REGION Network 15
   RUNG wire#powerrail
      { S7_Templates := "SrcType := Int" } EQ_Contact(in1 := "DB_general".Piston_2_Cursa_Completa, in2 := 25)
      R_Coil( "DB_HMI".Viz_Platforma_Libera )
   END_RUNG
   // the same network as SCL:
   IF "DB_general".Piston_2_Cursa_Completa = 25 THEN "DB_HMI".Viz_Platforma_Libera := FALSE; END_IF;
END_REGION
END_FUNCTION_BLOCK

FUNCTION_BLOCK "Piston_Incarcare"   // FB19, LAD
{ S7_Optimized_Access := 'FALSE' }
VERSION : 0.1
   VAR_TEMP   // added for the SCL form of the ladder/FBD networks
      _w1 : Bool;
      _w2 : Bool;
      _w3 : Bool;
      _w4 : Bool;
      _w5 : Bool;
      _w6 : Bool;
      _w7 : Bool;
   END_VAR
BEGIN

REGION Network 1
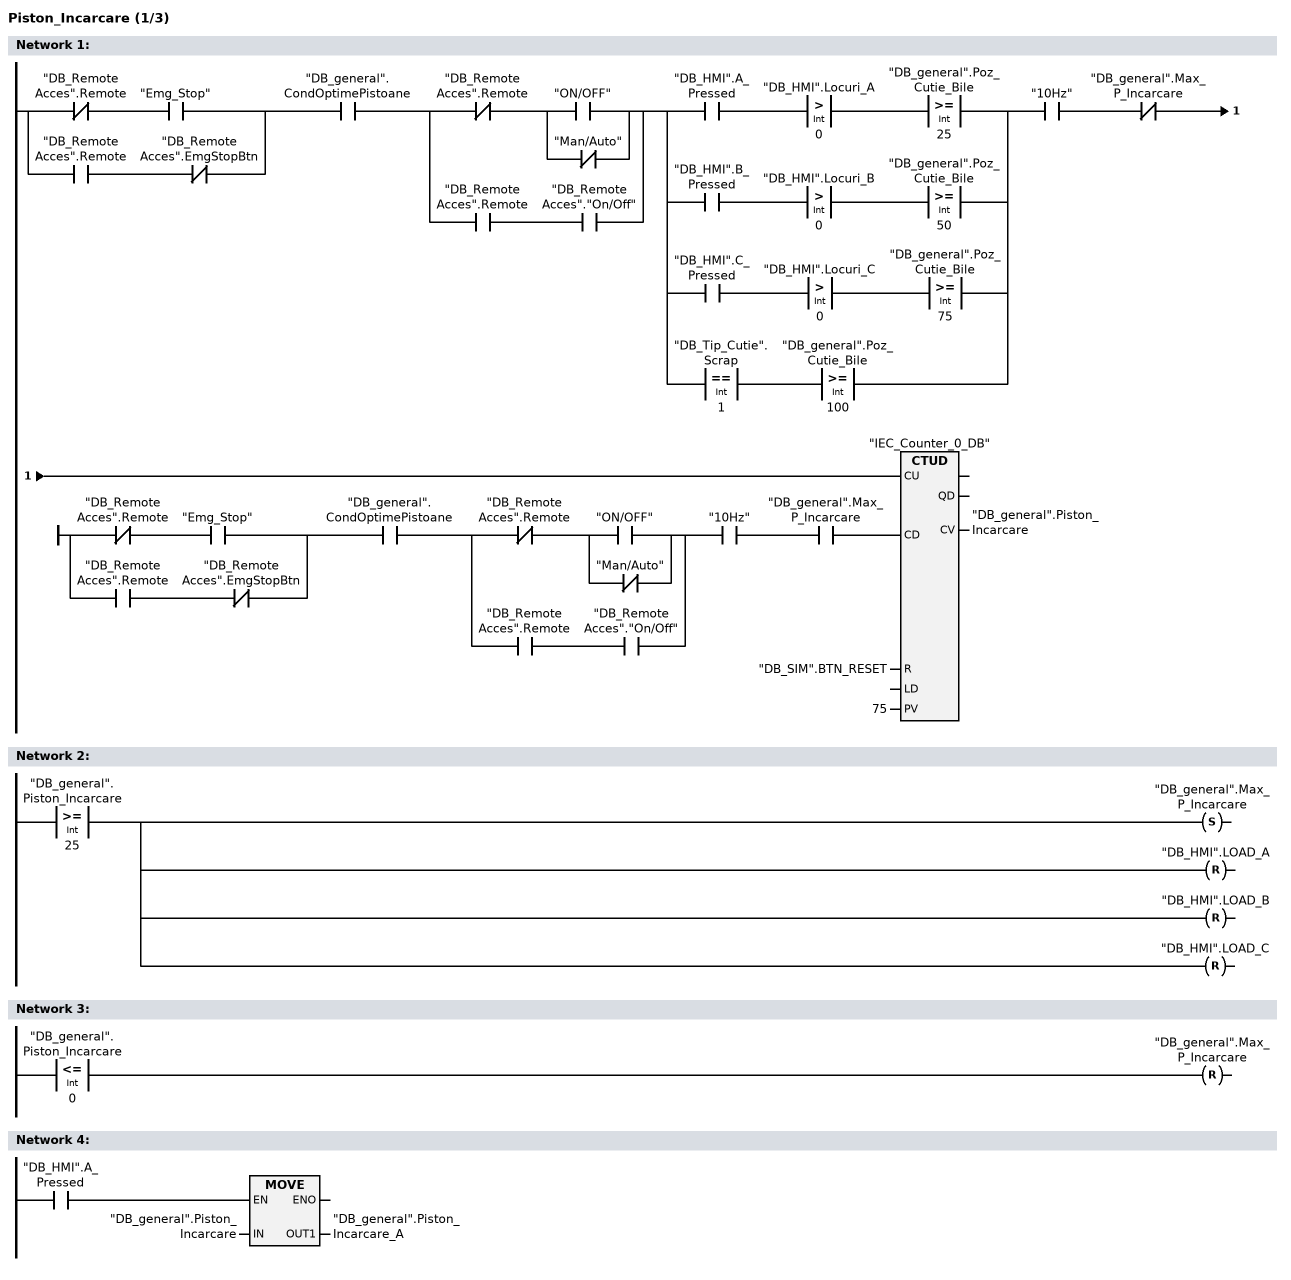
   "IEC_Counter_0_DB".CTUD(CU := ((NOT "DB_RemoteAcces".Remote AND "Emg_Stop") OR ("DB_RemoteAcces".Remote AND NOT "DB_RemoteAcces".EmgStopBtn)) AND "DB_general".CondOptimePistoane AND ((NOT "DB_RemoteAcces".Remote AND ("ON/OFF" OR NOT "Man/Auto")) OR ("DB_RemoteAcces".Remote AND "DB_RemoteAcces"."On/Off")) AND (("DB_HMI".A_Pressed AND ("DB_HMI".Locuri_A > 0) AND ("DB_general".Poz_Cutie_Bile >= 25)) OR ("DB_HMI".B_Pressed AND ("DB_HMI".Locuri_B > 0) AND ("DB_general".Poz_Cutie_Bile >= 50)) OR ("DB_HMI".C_Pressed AND ("DB_HMI".Locuri_C > 0) AND ("DB_general".Poz_Cutie_Bile >= 75)) OR (("DB_Tip_Cutie".Scrap = 1) AND ("DB_general".Poz_Cutie_Bile >= 100))) AND "10Hz" AND NOT "DB_general".Max_P_Incarcare,
                           CD := ((NOT "DB_RemoteAcces".Remote AND "Emg_Stop") OR ("DB_RemoteAcces".Remote AND NOT "DB_RemoteAcces".EmgStopBtn)) AND "DB_general".CondOptimePistoane AND ((NOT "DB_RemoteAcces".Remote AND ("ON/OFF" OR NOT "Man/Auto")) OR ("DB_RemoteAcces".Remote AND "DB_RemoteAcces"."On/Off")) AND "10Hz" AND "DB_general".Max_P_Incarcare,
                           R := "DB_SIM".BTN_RESET,
                           PV := 75,
                           CV => "DB_general".Piston_Incarcare);
END_REGION

REGION Network 2
   RUNG wire#powerrail
      { S7_Templates := "SrcType := Int" } GE_Contact(in1 := "DB_general".Piston_Incarcare, in2 := 25)
      wire#w1
      S_Coil( "DB_general".Max_P_Incarcare )
   END_RUNG
   RUNG wire#w1
      R_Coil( "DB_HMI".LOAD_A )
   END_RUNG
   RUNG wire#w1
      R_Coil( "DB_HMI".LOAD_B )
   END_RUNG
   RUNG wire#w1
      R_Coil( "DB_HMI".LOAD_C )
   END_RUNG
   // the same network as SCL:
   IF "DB_general".Piston_Incarcare >= 25 THEN
       "DB_general".Max_P_Incarcare := TRUE;
       "DB_HMI".LOAD_A := FALSE;
       "DB_HMI".LOAD_B := FALSE;
       "DB_HMI".LOAD_C := FALSE;
   END_IF;
END_REGION

REGION Network 3
   RUNG wire#powerrail
      { S7_Templates := "SrcType := Int" } LE_Contact(in1 := "DB_general".Piston_Incarcare, in2 := 0)
      R_Coil( "DB_general".Max_P_Incarcare )
   END_RUNG
   // the same network as SCL:
   IF "DB_general".Piston_Incarcare <= 0 THEN "DB_general".Max_P_Incarcare := FALSE; END_IF;
END_REGION

REGION Network 4
   RUNG wire#powerrail
      Contact( "DB_HMI".A_Pressed )
      { S7_GenerateENO := "TRUE" } Move(in := "DB_general".Piston_Incarcare, out1 => "DB_general".Piston_Incarcare_A)
   END_RUNG
   // the same network as SCL:
   IF "DB_HMI".A_Pressed THEN "DB_general".Piston_Incarcare_A := "DB_general".Piston_Incarcare; END_IF;
END_REGION

REGION Network 5
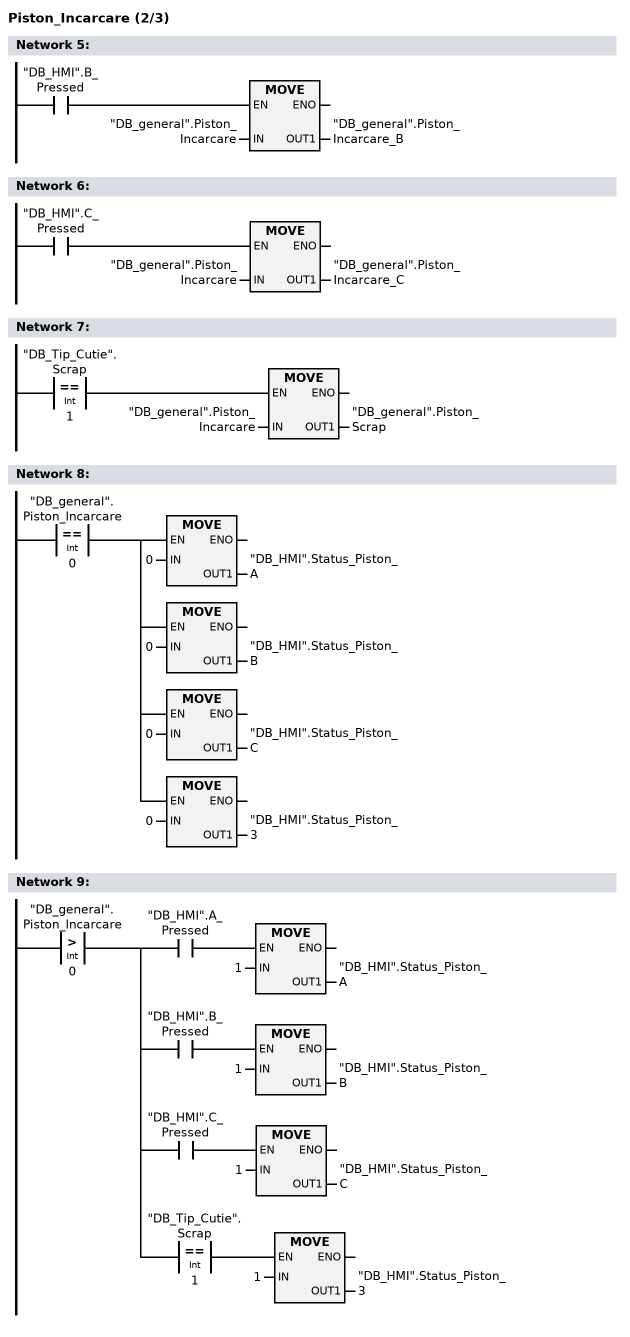
   RUNG wire#powerrail
      Contact( "DB_HMI".B_Pressed )
      { S7_GenerateENO := "TRUE" } Move(in := "DB_general".Piston_Incarcare, out1 => "DB_general".Piston_Incarcare_B)
   END_RUNG
   // the same network as SCL:
   IF "DB_HMI".B_Pressed THEN "DB_general".Piston_Incarcare_B := "DB_general".Piston_Incarcare; END_IF;
END_REGION

REGION Network 6
   RUNG wire#powerrail
      Contact( "DB_HMI".C_Pressed )
      { S7_GenerateENO := "TRUE" } Move(in := "DB_general".Piston_Incarcare, out1 => "DB_general".Piston_Incarcare_C)
   END_RUNG
   // the same network as SCL:
   IF "DB_HMI".C_Pressed THEN "DB_general".Piston_Incarcare_C := "DB_general".Piston_Incarcare; END_IF;
END_REGION

REGION Network 7
   RUNG wire#powerrail
      { S7_Templates := "SrcType := Int" } EQ_Contact(in1 := "DB_Tip_Cutie".Scrap, in2 := 1)
      { S7_GenerateENO := "TRUE" } Move(in := "DB_general".Piston_Incarcare, out1 => "DB_general".Piston_Scrap)
   END_RUNG
   // the same network as SCL:
   IF "DB_Tip_Cutie".Scrap = 1 THEN "DB_general".Piston_Scrap := "DB_general".Piston_Incarcare; END_IF;
END_REGION

REGION Network 8
   RUNG wire#powerrail
      { S7_Templates := "SrcType := Int" } EQ_Contact(in1 := "DB_general".Piston_Incarcare, in2 := 0)
      wire#w1
      { S7_GenerateENO := "TRUE" } Move(in := 0, out1 => "DB_HMI".Status_Piston_A)
   END_RUNG
   RUNG wire#w1
      { S7_GenerateENO := "TRUE" } Move(in := 0, out1 => "DB_HMI".Status_Piston_B)
   END_RUNG
   RUNG wire#w1
      { S7_GenerateENO := "TRUE" } Move(in := 0, out1 => "DB_HMI".Status_Piston_C)
   END_RUNG
   RUNG wire#w1
      { S7_GenerateENO := "TRUE" } Move(in := 0, out1 => "DB_HMI".Status_Piston_3)
   END_RUNG
   // the same network as SCL:
   IF "DB_general".Piston_Incarcare = 0 THEN
       "DB_HMI".Status_Piston_A := 0;
       "DB_HMI".Status_Piston_B := 0;
       "DB_HMI".Status_Piston_C := 0;
       "DB_HMI".Status_Piston_3 := 0;
   END_IF;
END_REGION

REGION Network 9
   RUNG wire#powerrail
      { S7_Templates := "SrcType := Int" } GT_Contact(in1 := "DB_general".Piston_Incarcare, in2 := 0)
      wire#w1
      Contact( "DB_HMI".A_Pressed )
      { S7_GenerateENO := "TRUE" } Move(in := 1, out1 => "DB_HMI".Status_Piston_A)
   END_RUNG
   RUNG wire#w1
      Contact( "DB_HMI".B_Pressed )
      { S7_GenerateENO := "TRUE" } Move(in := 1, out1 => "DB_HMI".Status_Piston_B)
   END_RUNG
   RUNG wire#w1
      Contact( "DB_HMI".C_Pressed )
      { S7_GenerateENO := "TRUE" } Move(in := 1, out1 => "DB_HMI".Status_Piston_C)
   END_RUNG
   RUNG wire#w1
      { S7_Templates := "SrcType := Int" } EQ_Contact(in1 := "DB_Tip_Cutie".Scrap, in2 := 1)
      { S7_GenerateENO := "TRUE" } Move(in := 1, out1 => "DB_HMI".Status_Piston_3)
   END_RUNG
   // the same network as SCL:
   #_w1 := "DB_general".Piston_Incarcare > 0;
   IF #_w1 AND "DB_HMI".A_Pressed THEN "DB_HMI".Status_Piston_A := 1; END_IF;
   IF #_w1 AND "DB_HMI".B_Pressed THEN "DB_HMI".Status_Piston_B := 1; END_IF;
   IF #_w1 AND "DB_HMI".C_Pressed THEN "DB_HMI".Status_Piston_C := 1; END_IF;
   IF #_w1 AND ("DB_Tip_Cutie".Scrap = 1) THEN "DB_HMI".Status_Piston_3 := 1; END_IF;
END_REGION

REGION Network 10
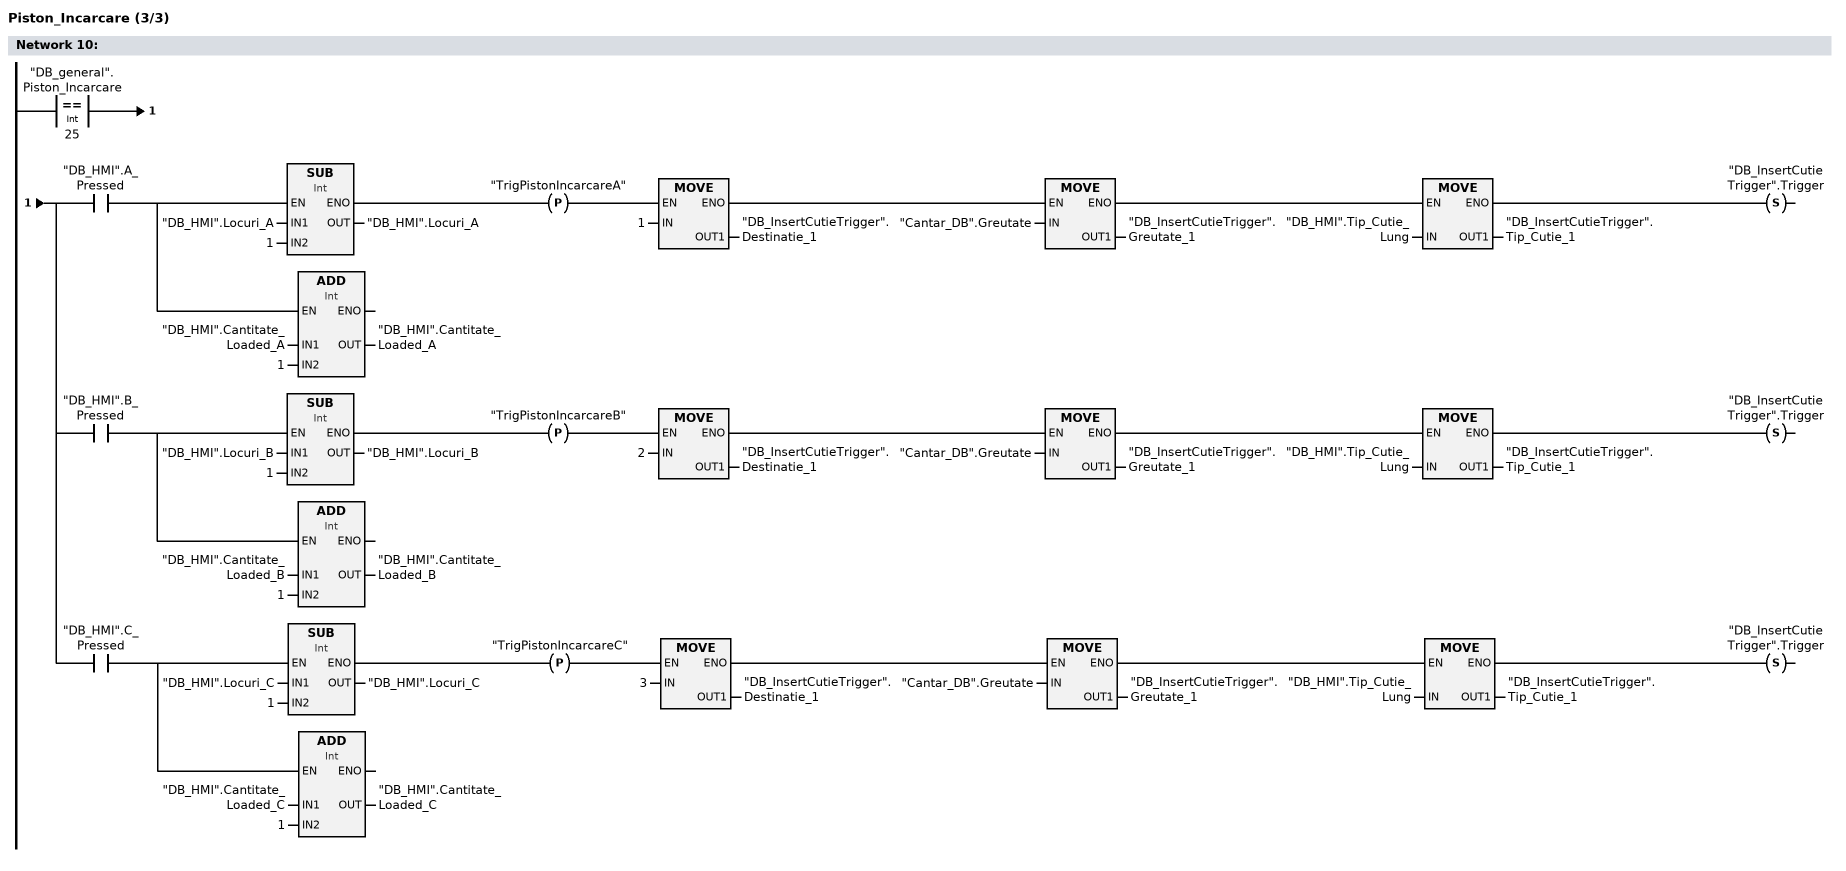
   RUNG wire#powerrail
      { S7_Templates := "SrcType := Int" } EQ_Contact(in1 := "DB_general".Piston_Incarcare, in2 := 25)
      wire#w1
      Contact( "DB_HMI".A_Pressed )
      wire#w2
      { S7_Templates := "SrcType := Int"; S7_GenerateENO := "TRUE" } Sub(in1 := "DB_HMI".Locuri_A, in2 := 1, out => "DB_HMI".Locuri_A)
      P_Trig( "TrigPistonIncarcareA" )
      { S7_GenerateENO := "TRUE" } Move(in := 1, out1 => "DB_InsertCutieTrigger".Destinatie_1)
      { S7_GenerateENO := "TRUE" } Move(in := "Cantar_DB".Greutate, out1 => "DB_InsertCutieTrigger".Greutate_1)
      { S7_GenerateENO := "TRUE" } Move(in := "DB_HMI".Tip_Cutie_Lung, out1 => "DB_InsertCutieTrigger".Tip_Cutie_1)
      S_Coil( "DB_InsertCutieTrigger".Trigger )
   END_RUNG
   RUNG wire#w2
      { S7_Templates := "SrcType := Int"; S7_GenerateENO := "TRUE" } Add(in1 := "DB_HMI".Cantitate_Loaded_A, in2 := 1, out => "DB_HMI".Cantitate_Loaded_A)
   END_RUNG
   RUNG wire#w1
      Contact( "DB_HMI".B_Pressed )
      wire#w3
      { S7_Templates := "SrcType := Int"; S7_GenerateENO := "TRUE" } Sub(in1 := "DB_HMI".Locuri_B, in2 := 1, out => "DB_HMI".Locuri_B)
      P_Trig( "TrigPistonIncarcareB" )
      { S7_GenerateENO := "TRUE" } Move(in := 2, out1 => "DB_InsertCutieTrigger".Destinatie_1)
      { S7_GenerateENO := "TRUE" } Move(in := "Cantar_DB".Greutate, out1 => "DB_InsertCutieTrigger".Greutate_1)
      { S7_GenerateENO := "TRUE" } Move(in := "DB_HMI".Tip_Cutie_Lung, out1 => "DB_InsertCutieTrigger".Tip_Cutie_1)
      S_Coil( "DB_InsertCutieTrigger".Trigger )
   END_RUNG
   RUNG wire#w3
      { S7_Templates := "SrcType := Int"; S7_GenerateENO := "TRUE" } Add(in1 := "DB_HMI".Cantitate_Loaded_B, in2 := 1, out => "DB_HMI".Cantitate_Loaded_B)
   END_RUNG
   RUNG wire#w1
      Contact( "DB_HMI".C_Pressed )
      wire#w4
      { S7_Templates := "SrcType := Int"; S7_GenerateENO := "TRUE" } Sub(in1 := "DB_HMI".Locuri_C, in2 := 1, out => "DB_HMI".Locuri_C)
      P_Trig( "TrigPistonIncarcareC" )
      { S7_GenerateENO := "TRUE" } Move(in := 3, out1 => "DB_InsertCutieTrigger".Destinatie_1)
      { S7_GenerateENO := "TRUE" } Move(in := "Cantar_DB".Greutate, out1 => "DB_InsertCutieTrigger".Greutate_1)
      { S7_GenerateENO := "TRUE" } Move(in := "DB_HMI".Tip_Cutie_Lung, out1 => "DB_InsertCutieTrigger".Tip_Cutie_1)
      S_Coil( "DB_InsertCutieTrigger".Trigger )
   END_RUNG
   RUNG wire#w4
      { S7_Templates := "SrcType := Int"; S7_GenerateENO := "TRUE" } Add(in1 := "DB_HMI".Cantitate_Loaded_C, in2 := 1, out => "DB_HMI".Cantitate_Loaded_C)
   END_RUNG
   // the same network as SCL:
   // ENO of a box is taken as its EN; it also drops when the box reports an error
   #_w1 := "DB_general".Piston_Incarcare = 25;
   #_w2 := #_w1 AND "DB_HMI".A_Pressed;
   IF #_w2 THEN "DB_HMI".Locuri_A := "DB_HMI".Locuri_A - 1; END_IF;
   #_w3 := #_w2 AND NOT "TrigPistonIncarcareA";   // rising edge
   "TrigPistonIncarcareA" := #_w2;
   IF #_w3 THEN
       "DB_InsertCutieTrigger".Destinatie_1 := 1;
       "DB_InsertCutieTrigger".Greutate_1 := "Cantar_DB".Greutate;
       "DB_InsertCutieTrigger".Tip_Cutie_1 := "DB_HMI".Tip_Cutie_Lung;
       "DB_InsertCutieTrigger".Trigger := TRUE;
   END_IF;
   IF #_w2 THEN "DB_HMI".Cantitate_Loaded_A := "DB_HMI".Cantitate_Loaded_A + 1; END_IF;
   #_w4 := #_w1 AND "DB_HMI".B_Pressed;
   IF #_w4 THEN "DB_HMI".Locuri_B := "DB_HMI".Locuri_B - 1; END_IF;
   #_w5 := #_w4 AND NOT "TrigPistonIncarcareB";   // rising edge
   "TrigPistonIncarcareB" := #_w4;
   IF #_w5 THEN
       "DB_InsertCutieTrigger".Destinatie_1 := 2;
       "DB_InsertCutieTrigger".Greutate_1 := "Cantar_DB".Greutate;
       "DB_InsertCutieTrigger".Tip_Cutie_1 := "DB_HMI".Tip_Cutie_Lung;
       "DB_InsertCutieTrigger".Trigger := TRUE;
   END_IF;
   IF #_w4 THEN "DB_HMI".Cantitate_Loaded_B := "DB_HMI".Cantitate_Loaded_B + 1; END_IF;
   #_w6 := #_w1 AND "DB_HMI".C_Pressed;
   IF #_w6 THEN "DB_HMI".Locuri_C := "DB_HMI".Locuri_C - 1; END_IF;
   #_w7 := #_w6 AND NOT "TrigPistonIncarcareC";   // rising edge
   "TrigPistonIncarcareC" := #_w6;
   IF #_w7 THEN
       "DB_InsertCutieTrigger".Destinatie_1 := 3;
       "DB_InsertCutieTrigger".Greutate_1 := "Cantar_DB".Greutate;
       "DB_InsertCutieTrigger".Tip_Cutie_1 := "DB_HMI".Tip_Cutie_Lung;
       "DB_InsertCutieTrigger".Trigger := TRUE;
   END_IF;
   IF #_w6 THEN "DB_HMI".Cantitate_Loaded_C := "DB_HMI".Cantitate_Loaded_C + 1; END_IF;
END_REGION
END_FUNCTION_BLOCK

FUNCTION "Vizibilitate_Platforme/Colete" : Void   // FC1, LAD
{ S7_Optimized_Access := 'FALSE' }
VERSION : 0.1
BEGIN

REGION Network 1: Caz A apasat setare vizibilitate / Sichtbarkeitseinstellung für Fall „A“.
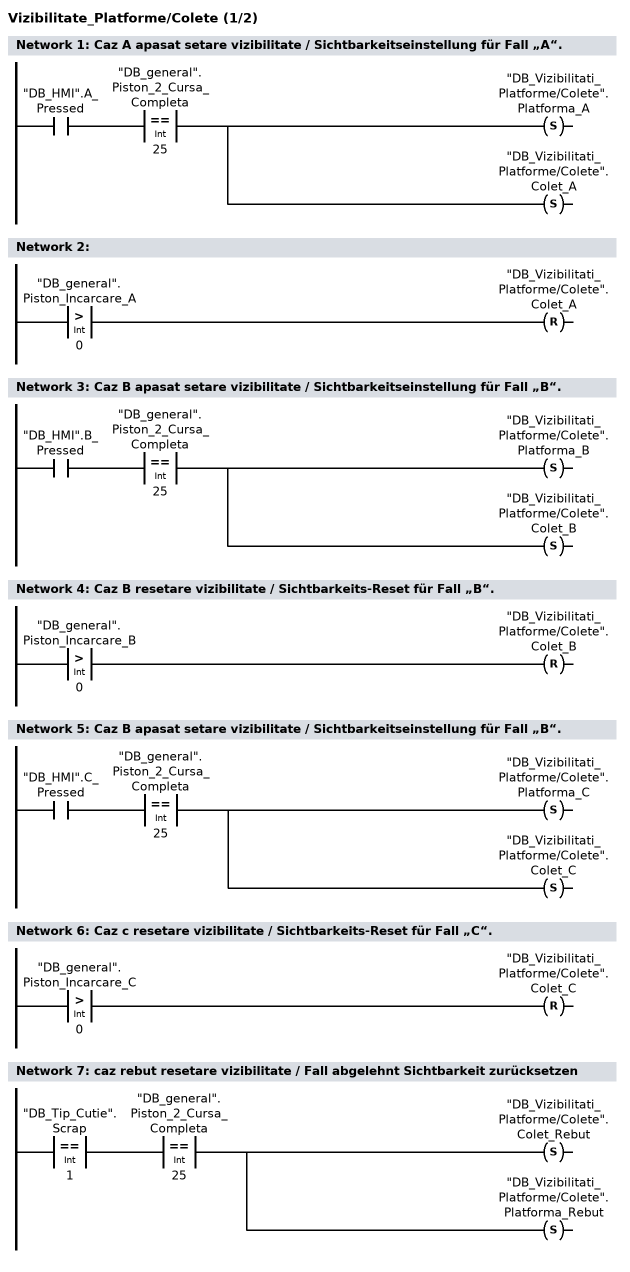
   RUNG wire#powerrail
      Contact( "DB_HMI".A_Pressed )
      { S7_Templates := "SrcType := Int" } EQ_Contact(in1 := "DB_general".Piston_2_Cursa_Completa, in2 := 25)
      wire#w1
      S_Coil( "DB_Vizibilitati_Platforme/Colete".Platforma_A )
   END_RUNG
   RUNG wire#w1
      S_Coil( "DB_Vizibilitati_Platforme/Colete".Colet_A )
   END_RUNG
   // the same network as SCL:
   IF "DB_HMI".A_Pressed AND ("DB_general".Piston_2_Cursa_Completa = 25) THEN
       "DB_Vizibilitati_Platforme/Colete".Platforma_A := TRUE;
       "DB_Vizibilitati_Platforme/Colete".Colet_A := TRUE;
   END_IF;
END_REGION

REGION Network 2
   RUNG wire#powerrail
      { S7_Templates := "SrcType := Int" } GT_Contact(in1 := "DB_general".Piston_Incarcare_A, in2 := 0)
      R_Coil( "DB_Vizibilitati_Platforme/Colete".Colet_A )
   END_RUNG
   // the same network as SCL:
   IF "DB_general".Piston_Incarcare_A > 0 THEN "DB_Vizibilitati_Platforme/Colete".Colet_A := FALSE; END_IF;
END_REGION

REGION Network 3: Caz B apasat setare vizibilitate / Sichtbarkeitseinstellung für Fall „B“.
   RUNG wire#powerrail
      Contact( "DB_HMI".B_Pressed )
      { S7_Templates := "SrcType := Int" } EQ_Contact(in1 := "DB_general".Piston_2_Cursa_Completa, in2 := 25)
      wire#w1
      S_Coil( "DB_Vizibilitati_Platforme/Colete".Platforma_B )
   END_RUNG
   RUNG wire#w1
      S_Coil( "DB_Vizibilitati_Platforme/Colete".Colet_B )
   END_RUNG
   // the same network as SCL:
   IF "DB_HMI".B_Pressed AND ("DB_general".Piston_2_Cursa_Completa = 25) THEN
       "DB_Vizibilitati_Platforme/Colete".Platforma_B := TRUE;
       "DB_Vizibilitati_Platforme/Colete".Colet_B := TRUE;
   END_IF;
END_REGION

REGION Network 4: Caz B resetare vizibilitate / Sichtbarkeits-Reset für Fall „B“.
   RUNG wire#powerrail
      { S7_Templates := "SrcType := Int" } GT_Contact(in1 := "DB_general".Piston_Incarcare_B, in2 := 0)
      R_Coil( "DB_Vizibilitati_Platforme/Colete".Colet_B )
   END_RUNG
   // the same network as SCL:
   IF "DB_general".Piston_Incarcare_B > 0 THEN "DB_Vizibilitati_Platforme/Colete".Colet_B := FALSE; END_IF;
END_REGION

REGION Network 5: Caz B apasat setare vizibilitate / Sichtbarkeitseinstellung für Fall „B“.
   RUNG wire#powerrail
      Contact( "DB_HMI".C_Pressed )
      { S7_Templates := "SrcType := Int" } EQ_Contact(in1 := "DB_general".Piston_2_Cursa_Completa, in2 := 25)
      wire#w1
      S_Coil( "DB_Vizibilitati_Platforme/Colete".Platforma_C )
   END_RUNG
   RUNG wire#w1
      S_Coil( "DB_Vizibilitati_Platforme/Colete".Colet_C )
   END_RUNG
   // the same network as SCL:
   IF "DB_HMI".C_Pressed AND ("DB_general".Piston_2_Cursa_Completa = 25) THEN
       "DB_Vizibilitati_Platforme/Colete".Platforma_C := TRUE;
       "DB_Vizibilitati_Platforme/Colete".Colet_C := TRUE;
   END_IF;
END_REGION

REGION Network 6: Caz c resetare vizibilitate / Sichtbarkeits-Reset für Fall „C“.
   RUNG wire#powerrail
      { S7_Templates := "SrcType := Int" } GT_Contact(in1 := "DB_general".Piston_Incarcare_C, in2 := 0)
      R_Coil( "DB_Vizibilitati_Platforme/Colete".Colet_C )
   END_RUNG
   // the same network as SCL:
   IF "DB_general".Piston_Incarcare_C > 0 THEN "DB_Vizibilitati_Platforme/Colete".Colet_C := FALSE; END_IF;
END_REGION

REGION Network 7: caz rebut resetare vizibilitate / Fall abgelehnt Sichtbarkeit zurücksetzen
   RUNG wire#powerrail
      { S7_Templates := "SrcType := Int" } EQ_Contact(in1 := "DB_Tip_Cutie".Scrap, in2 := 1)
      { S7_Templates := "SrcType := Int" } EQ_Contact(in1 := "DB_general".Piston_2_Cursa_Completa, in2 := 25)
      wire#w1
      S_Coil( "DB_Vizibilitati_Platforme/Colete".Colet_Rebut )
   END_RUNG
   RUNG wire#w1
      S_Coil( "DB_Vizibilitati_Platforme/Colete".Platforma_Rebut )
   END_RUNG
   // the same network as SCL:
   IF ("DB_Tip_Cutie".Scrap = 1) AND ("DB_general".Piston_2_Cursa_Completa = 25) THEN
       "DB_Vizibilitati_Platforme/Colete".Colet_Rebut := TRUE;
       "DB_Vizibilitati_Platforme/Colete".Platforma_Rebut := TRUE;
   END_IF;
END_REGION

REGION Network 8
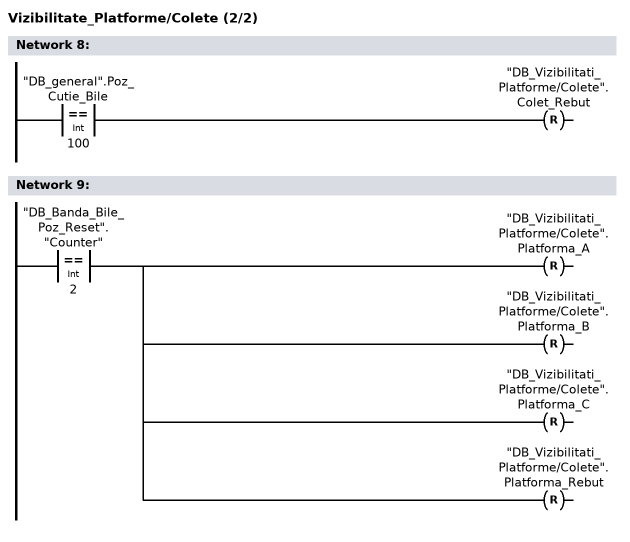
   RUNG wire#powerrail
      { S7_Templates := "SrcType := Int" } EQ_Contact(in1 := "DB_general".Poz_Cutie_Bile, in2 := 100)
      R_Coil( "DB_Vizibilitati_Platforme/Colete".Colet_Rebut )
   END_RUNG
   // the same network as SCL:
   IF "DB_general".Poz_Cutie_Bile = 100 THEN "DB_Vizibilitati_Platforme/Colete".Colet_Rebut := FALSE; END_IF;
END_REGION

REGION Network 9
   RUNG wire#powerrail
      { S7_Templates := "SrcType := Int" } EQ_Contact(in1 := "DB_Banda_Bile_Poz_Reset"."Counter", in2 := 2)
      wire#w1
      R_Coil( "DB_Vizibilitati_Platforme/Colete".Platforma_A )
   END_RUNG
   RUNG wire#w1
      R_Coil( "DB_Vizibilitati_Platforme/Colete".Platforma_B )
   END_RUNG
   RUNG wire#w1
      R_Coil( "DB_Vizibilitati_Platforme/Colete".Platforma_C )
   END_RUNG
   RUNG wire#w1
      R_Coil( "DB_Vizibilitati_Platforme/Colete".Platforma_Rebut )
   END_RUNG
   // the same network as SCL:
   IF "DB_Banda_Bile_Poz_Reset"."Counter" = 2 THEN
       "DB_Vizibilitati_Platforme/Colete".Platforma_A := FALSE;
       "DB_Vizibilitati_Platforme/Colete".Platforma_B := FALSE;
       "DB_Vizibilitati_Platforme/Colete".Platforma_C := FALSE;
       "DB_Vizibilitati_Platforme/Colete".Platforma_Rebut := FALSE;
   END_IF;
END_REGION
END_FUNCTION

// folder: Statie Incarcare/Functii

FUNCTION_BLOCK "Banda_Bile"   // FB16, SCL
{ S7_Optimized_Access := 'FALSE' }
VERSION : 0.1
   VAR_INPUT
      "Man/Auto" : Bool;
      BTN_Transport : Bool;
      Poz_Cutie_1 : Int;
      Emg_Stop : Bool;
      Btn_A : Bool;
      Btn_B : Bool;
      Btn_C : Bool;
   END_VAR
   VAR_OUTPUT
      Status_Banda_Bile : Bool;
   END_VAR
   VAR
      Btn_Transport_Pressed : Bool;
   END_VAR
BEGIN
   //IF #BTN_Transport THEN
     //  #Btn_Transport_Pressed := true;

   //END_IF;



       IF #Poz_Cutie_1 >48 AND "DB_HMI".Transport AND "DB_general".Piston_2_Cursa_Completa =0 AND (#Btn_A OR #Btn_B OR #Btn_C OR "DB_Tip_Cutie".Scrap = 1) THEN

           #Status_Banda_Bile := TRUE;
       ELSE
           #Status_Banda_Bile := FALSE;
           #Btn_Transport_Pressed := FALSE;


       END_IF;
END_FUNCTION_BLOCK

FUNCTION "Banda_Bile_Poz_Reset" : Void   // FC9, LAD
{ S7_Optimized_Access := 'FALSE' }
VERSION : 0.1
BEGIN

REGION Network 1
   // Atunci cand platforma cu bile trece de doua ori prin dreptul unui punct inseamna ca s a efectuat descarcarea si ca op ar trebui sa introduca o alta destinatie
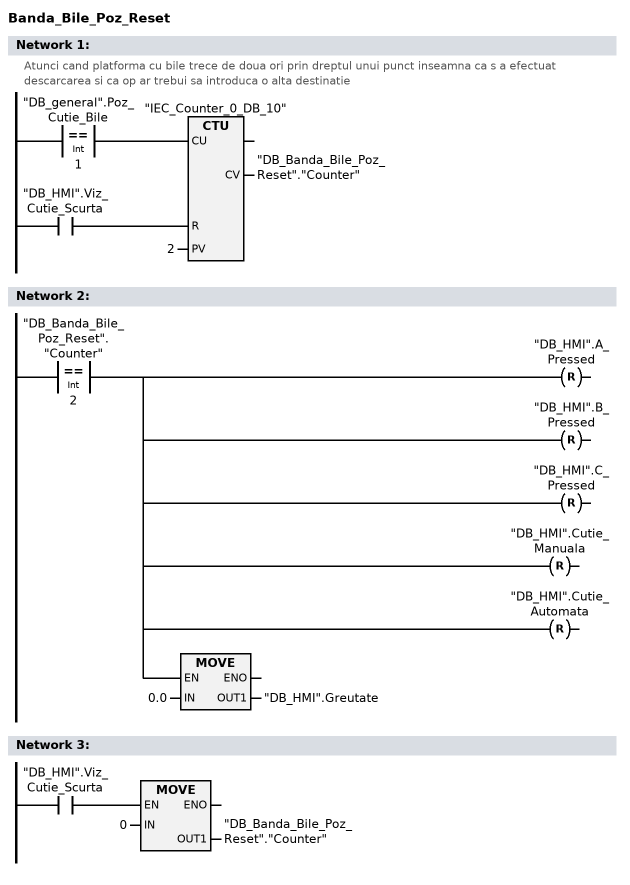
   "IEC_Counter_0_DB_10".CTU(CU := "DB_general".Poz_Cutie_Bile = 1,
                           R := "DB_HMI".Viz_Cutie_Scurta,
                           PV := 2,
                           CV => "DB_Banda_Bile_Poz_Reset"."Counter");
END_REGION

REGION Network 2
   RUNG wire#powerrail
      { S7_Templates := "SrcType := Int" } EQ_Contact(in1 := "DB_Banda_Bile_Poz_Reset"."Counter", in2 := 2)
      wire#w1
      R_Coil( "DB_HMI".A_Pressed )
   END_RUNG
   RUNG wire#w1
      R_Coil( "DB_HMI".B_Pressed )
   END_RUNG
   RUNG wire#w1
      R_Coil( "DB_HMI".C_Pressed )
   END_RUNG
   RUNG wire#w1
      R_Coil( "DB_HMI".Cutie_Manuala )
   END_RUNG
   RUNG wire#w1
      R_Coil( "DB_HMI".Cutie_Automata )
   END_RUNG
   RUNG wire#w1
      { S7_GenerateENO := "TRUE" } Move(in := 0.0, out1 => "DB_HMI".Greutate)
   END_RUNG
   // the same network as SCL:
   IF "DB_Banda_Bile_Poz_Reset"."Counter" = 2 THEN
       "DB_HMI".A_Pressed := FALSE;
       "DB_HMI".B_Pressed := FALSE;
       "DB_HMI".C_Pressed := FALSE;
       "DB_HMI".Cutie_Manuala := FALSE;
       "DB_HMI".Cutie_Automata := FALSE;
       "DB_HMI".Greutate := 0.0;
   END_IF;
END_REGION

REGION Network 3
   RUNG wire#powerrail
      Contact( "DB_HMI".Viz_Cutie_Scurta )
      { S7_GenerateENO := "TRUE" } Move(in := 0, out1 => "DB_Banda_Bile_Poz_Reset"."Counter")
   END_RUNG
   // the same network as SCL:
   IF "DB_HMI".Viz_Cutie_Scurta THEN "DB_Banda_Bile_Poz_Reset"."Counter" := 0; END_IF;
END_REGION
END_FUNCTION

FUNCTION "GreutateTotala" : Void   // FC14, LAD
{ S7_Optimized_Access := 'FALSE' }
VERSION : 0.1
BEGIN

REGION Network 1
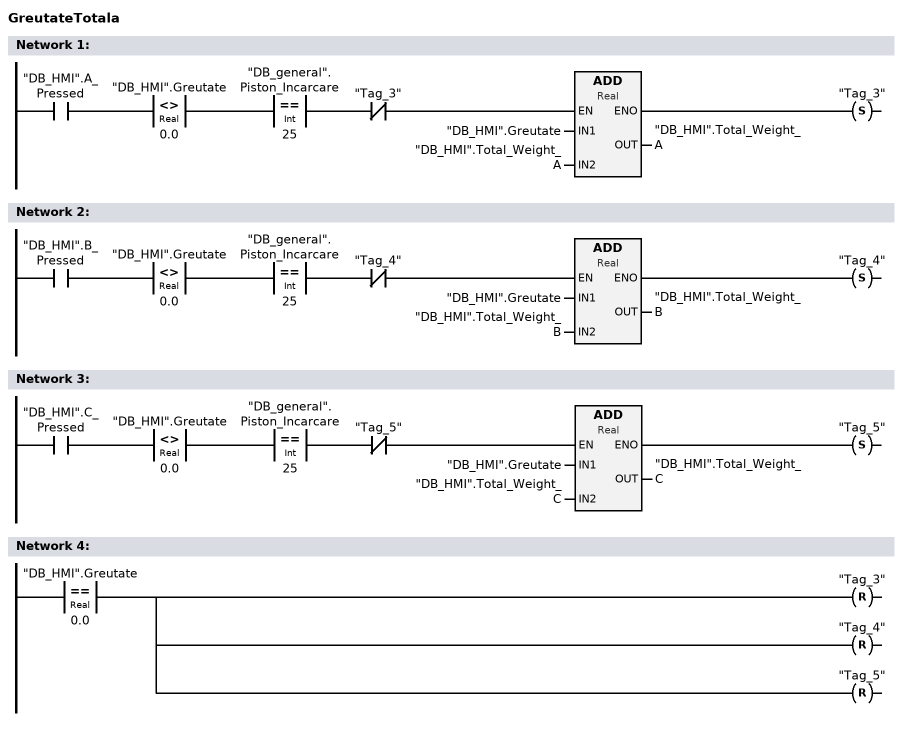
   RUNG wire#powerrail
      Contact( "DB_HMI".A_Pressed )
      { S7_Templates := "SrcType := Real" } NE_Contact(in1 := "DB_HMI".Greutate, in2 := 0.0)
      { S7_Templates := "SrcType := Int" } EQ_Contact(in1 := "DB_general".Piston_Incarcare, in2 := 25)
      I_Contact( "Tag_3" )
      { S7_Templates := "SrcType := Real"; S7_GenerateENO := "TRUE" } Add(in1 := "DB_HMI".Greutate, in2 := "DB_HMI".Total_Weight_A, out => "DB_HMI".Total_Weight_A)
      S_Coil( "Tag_3" )
   END_RUNG
   // the same network as SCL:
   // ENO of a box is taken as its EN; it also drops when the box reports an error
   IF "DB_HMI".A_Pressed AND ("DB_HMI".Greutate <> 0.0) AND ("DB_general".Piston_Incarcare = 25) AND NOT "Tag_3" THEN
       "DB_HMI".Total_Weight_A := "DB_HMI".Greutate + "DB_HMI".Total_Weight_A;
       "Tag_3" := TRUE;
   END_IF;
END_REGION

REGION Network 2
   RUNG wire#powerrail
      Contact( "DB_HMI".B_Pressed )
      { S7_Templates := "SrcType := Real" } NE_Contact(in1 := "DB_HMI".Greutate, in2 := 0.0)
      { S7_Templates := "SrcType := Int" } EQ_Contact(in1 := "DB_general".Piston_Incarcare, in2 := 25)
      I_Contact( "Tag_4" )
      { S7_Templates := "SrcType := Real"; S7_GenerateENO := "TRUE" } Add(in1 := "DB_HMI".Greutate, in2 := "DB_HMI".Total_Weight_B, out => "DB_HMI".Total_Weight_B)
      S_Coil( "Tag_4" )
   END_RUNG
   // the same network as SCL:
   // ENO of a box is taken as its EN; it also drops when the box reports an error
   IF "DB_HMI".B_Pressed AND ("DB_HMI".Greutate <> 0.0) AND ("DB_general".Piston_Incarcare = 25) AND NOT "Tag_4" THEN
       "DB_HMI".Total_Weight_B := "DB_HMI".Greutate + "DB_HMI".Total_Weight_B;
       "Tag_4" := TRUE;
   END_IF;
END_REGION

REGION Network 3
   RUNG wire#powerrail
      Contact( "DB_HMI".C_Pressed )
      { S7_Templates := "SrcType := Real" } NE_Contact(in1 := "DB_HMI".Greutate, in2 := 0.0)
      { S7_Templates := "SrcType := Int" } EQ_Contact(in1 := "DB_general".Piston_Incarcare, in2 := 25)
      I_Contact( "Tag_5" )
      { S7_Templates := "SrcType := Real"; S7_GenerateENO := "TRUE" } Add(in1 := "DB_HMI".Greutate, in2 := "DB_HMI".Total_Weight_C, out => "DB_HMI".Total_Weight_C)
      S_Coil( "Tag_5" )
   END_RUNG
   // the same network as SCL:
   // ENO of a box is taken as its EN; it also drops when the box reports an error
   IF "DB_HMI".C_Pressed AND ("DB_HMI".Greutate <> 0.0) AND ("DB_general".Piston_Incarcare = 25) AND NOT "Tag_5" THEN
       "DB_HMI".Total_Weight_C := "DB_HMI".Greutate + "DB_HMI".Total_Weight_C;
       "Tag_5" := TRUE;
   END_IF;
END_REGION

REGION Network 4
   RUNG wire#powerrail
      { S7_Templates := "SrcType := Real" } EQ_Contact(in1 := "DB_HMI".Greutate, in2 := 0.0)
      wire#w1
      R_Coil( "Tag_3" )
   END_RUNG
   RUNG wire#w1
      R_Coil( "Tag_4" )
   END_RUNG
   RUNG wire#w1
      R_Coil( "Tag_5" )
   END_RUNG
   // the same network as SCL:
   IF "DB_HMI".Greutate = 0.0 THEN
       "Tag_3" := FALSE;
       "Tag_4" := FALSE;
       "Tag_5" := FALSE;
   END_IF;
END_REGION
END_FUNCTION

// folder: Statie Retur

FUNCTION "BandaRetur" : Void   // FC20, LAD
{ S7_Optimized_Access := 'FALSE' }
VERSION : 0.1
BEGIN

REGION Network 1
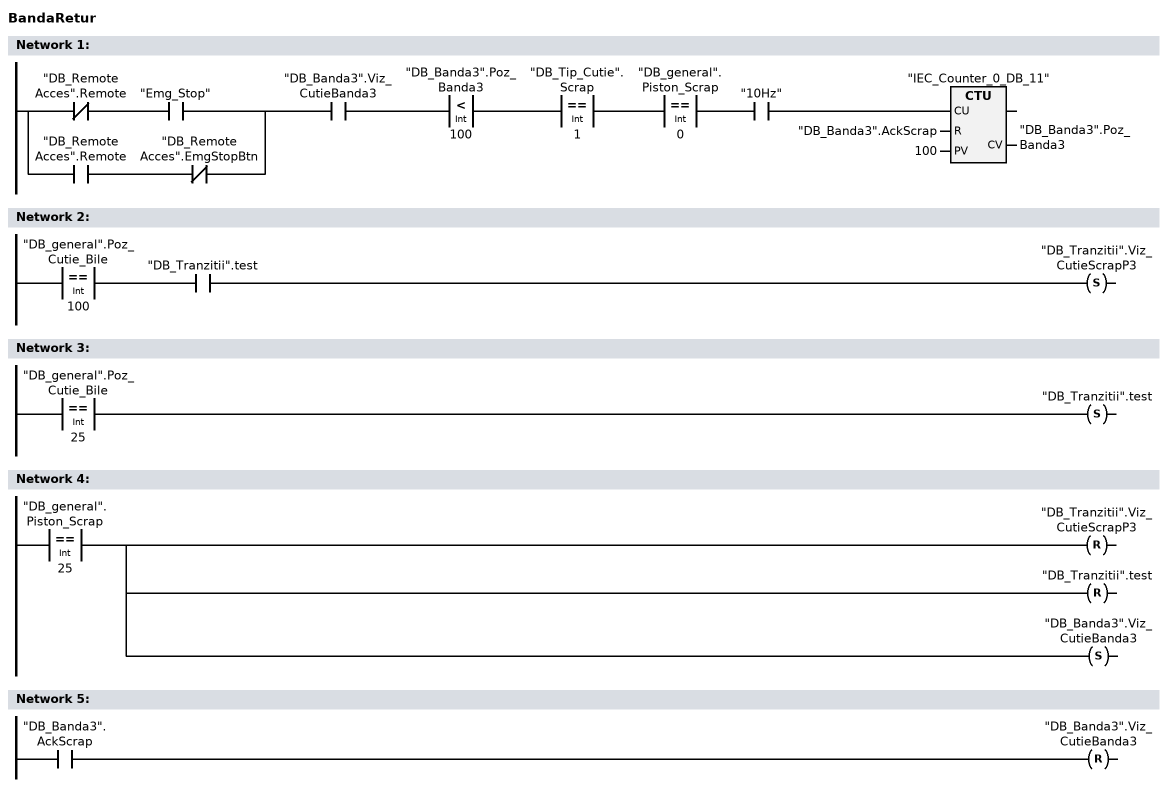
   "IEC_Counter_0_DB_11".CTU(CU := ((NOT "DB_RemoteAcces".Remote AND "Emg_Stop") OR ("DB_RemoteAcces".Remote AND NOT "DB_RemoteAcces".EmgStopBtn)) AND "DB_Banda3".Viz_CutieBanda3 AND ("DB_Banda3".Poz_Banda3 < 100) AND ("DB_Tip_Cutie".Scrap = 1) AND ("DB_general".Piston_Scrap = 0) AND "10Hz",
                           R := "DB_Banda3".AckScrap,
                           PV := 100,
                           CV => "DB_Banda3".Poz_Banda3);
END_REGION

REGION Network 2
   RUNG wire#powerrail
      { S7_Templates := "SrcType := Int" } EQ_Contact(in1 := "DB_general".Poz_Cutie_Bile, in2 := 100)
      Contact( "DB_Tranzitii".test )
      S_Coil( "DB_Tranzitii".Viz_CutieScrapP3 )
   END_RUNG
   // the same network as SCL:
   IF ("DB_general".Poz_Cutie_Bile = 100) AND "DB_Tranzitii".test THEN
       "DB_Tranzitii".Viz_CutieScrapP3 := TRUE;
   END_IF;
END_REGION

REGION Network 3
   RUNG wire#powerrail
      { S7_Templates := "SrcType := Int" } EQ_Contact(in1 := "DB_general".Poz_Cutie_Bile, in2 := 25)
      S_Coil( "DB_Tranzitii".test )
   END_RUNG
   // the same network as SCL:
   IF "DB_general".Poz_Cutie_Bile = 25 THEN "DB_Tranzitii".test := TRUE; END_IF;
END_REGION

REGION Network 4
   RUNG wire#powerrail
      { S7_Templates := "SrcType := Int" } EQ_Contact(in1 := "DB_general".Piston_Scrap, in2 := 25)
      wire#w1
      R_Coil( "DB_Tranzitii".Viz_CutieScrapP3 )
   END_RUNG
   RUNG wire#w1
      R_Coil( "DB_Tranzitii".test )
   END_RUNG
   RUNG wire#w1
      S_Coil( "DB_Banda3".Viz_CutieBanda3 )
   END_RUNG
   // the same network as SCL:
   IF "DB_general".Piston_Scrap = 25 THEN
       "DB_Tranzitii".Viz_CutieScrapP3 := FALSE;
       "DB_Tranzitii".test := FALSE;
       "DB_Banda3".Viz_CutieBanda3 := TRUE;
   END_IF;
END_REGION

REGION Network 5
   RUNG wire#powerrail
      Contact( "DB_Banda3".AckScrap )
      R_Coil( "DB_Banda3".Viz_CutieBanda3 )
   END_RUNG
   // the same network as SCL:
   IF "DB_Banda3".AckScrap THEN "DB_Banda3".Viz_CutieBanda3 := FALSE; END_IF;
END_REGION
END_FUNCTION

// ===== PLC "PLC_2"  CPU 1518-4 PN/DP =====

DATA_BLOCK "fb_DB"   // DB1
{ S7_Optimized_Access := 'TRUE' }
VERSION : 0.1
// stored: InstanceOfName fb
"fb"
BEGIN
END_DATA_BLOCK

FUNCTION_BLOCK "fb"   // FB1, GRAPH_PLUS
{ S7_Optimized_Access := 'TRUE' }
VERSION : 0.1
   VAR_INPUT
      OFF_SQ : Bool := false;   // Turn sequence off
      INIT_SQ : Bool := false;   // Set sequence to initial state
      ACK_EF : Bool := false;   // Acknowledge all errors and faults
      S_PREV : Bool := false;   // Output previous step in parameter S_NO
      S_NEXT : Bool := false;   // Indicate next step in parameter S_NO
      SW_AUTO : Bool := false;   // Automatic mode
      SW_TAP : Bool := false;   // Semiautomatic/switch with transition
      SW_TOP : Bool := false;   // Semiautomatic/ignore transition
      SW_MAN : Bool := false;   // Manual mode
      S_SEL : Int := 0;   // Select step to be output to S_NO
      S_ON : Bool := false;   // Activate step indicated in S_NO
      S_OFF : Bool := false;   // Deactivate step indicated S_NO
      T_PUSH : Bool := false;   // Enable transition to switch in semi automatic mode
   END_VAR
   VAR_OUTPUT
      S_NO : Int := 0;   // Step number
      S_MORE : Bool := false;   // More steps are available and can be shown in S_NO
      S_ACTIVE : Bool := false;   // Step indicated in S_NO is active
      ERR_FLT : Bool := false;   // Interlock or supervision group error
      AUTO_ON : Bool := false;   // Automatic mode is active
      TAP_ON : Bool := false;   // Semiautomatic mode/step with transition enabled
      TOP_ON : Bool := false;   // Semiautomatic mode/ignore transition enabled
      MAN_ON : Bool := false;   // Manual mode is active
   END_VAR
   VAR
      HMI_INFO : Array[0..8] of UInt;
      IF_PAR : G7_IfParPlus_V6;
      RT_DATA : G7_RTDataPlus_V6;   // Internal data area
      Trans1 : G7_TransitionPlus_V6;   // Transition structure
      Step1 : G7_StepPlus_V6;   // Step structure
      SINI : Array[0..1] of USInt;
      LSTT : Array[0..0] of USInt;
      ATAJ : Array[0..0] of USInt;
      ATAB : Array[0..0] of USInt;
      PSTT : Array[0..0] of USInt;
      NSTT : Array[0..0] of USInt;
      ASSJ : Array[0..0] of USInt;
      ASSB : Array[0..0] of USInt;
      PTTS : Array[0..0] of USInt;
      NTTS : Array[0..0] of USInt;
      SW_SQTS : Array[0..0] of USInt;
      SWITCH : Array[0..0] of USInt;
      TVX : Array[0..1] of USInt;
      TTX : Array[0..1] of USInt;
      TSX : Array[0..1] of USInt;
      S00X : Array[0..1] of USInt;
      SOFFX : Array[0..1] of USInt;
      SONX : Array[0..1] of USInt;
      SAX : Array[0..1] of USInt;
      SERRX : Array[0..1] of USInt;
      SMX : Array[0..1] of USInt;
      S0X : Array[0..1] of USInt;
      S1X : Array[0..1] of USInt;
      IL_ALARM_INST : Diag_Alarm;
      SUP_ALARM_INST : Diag_Alarm;
      STEP_TIME_ALARM_INST : Diag_Alarm;
      IEC_TIMER_INST : IEC_TIMER;
      TRANSACTION_FLAG : Bool := false;
   END_VAR
   // SINI[0] := 2;
   // PTTS[0] := 255;
   // TVX[0] := 16#1;
   // TTX[0] := 16#1;
   // TSX[0] := 16#1;
   // S00X[0] := 16#1;
   // SOFFX[0] := 16#1;
   // SONX[0] := 16#1;
   // SAX[0] := 16#1;
   // SERRX[0] := 16#1;
   // SMX[0] := 16#1;
   // S0X[0] := 16#1;
   // S1X[0] := 16#1;
BEGIN
